REGION Network 256
   RUNG wire#powerrail
      Contact( "EMS".Carrier[41].SDC_OUT.Faults.MotionOnFault )
      Coil( "Carrier_41_Motion_On_Fault" )
   END_RUNG
   // the same network as SCL:
   "Carrier_41_Motion_On_Fault" := "EMS".Carrier[41].SDC_OUT.Faults.MotionOnFault;
END_REGION

REGION Network 257
   RUNG wire#powerrail
      Contact( "EMS".Carrier[41].SDC_OUT.Faults.MotionOffFault )
      Coil( "Carrier_41_Motion_Off_Fault" )
   END_RUNG
   // the same network as SCL:
   "Carrier_41_Motion_Off_Fault" := "EMS".Carrier[41].SDC_OUT.Faults.MotionOffFault;
END_REGION

REGION Network 258
   RUNG wire#powerrail
      Contact( "EMS".Carrier[41].SDC_OUT.Faults.CarrierSpacingFault )
      Coil( "Carrier_41_Carrier_Spacing_Fault" )
   END_RUNG
   // the same network as SCL:
   "Carrier_41_Carrier_Spacing_Fault" := "EMS".Carrier[41].SDC_OUT.Faults.CarrierSpacingFault;
END_REGION

REGION Network 259
   RUNG wire#powerrail
      Move(in := "EMS".Carrier[42].SDC_OUT.Zone, out1 => "Carrier_42_Carrier_In_Zone")
   END_RUNG
   // the same network as SCL:
   "Carrier_42_Carrier_In_Zone" := "EMS".Carrier[42].SDC_OUT.Zone;
END_REGION

REGION Network 260
   RUNG wire#powerrail
      Move(in := "EMS".Carrier[42].SDC_OUT.CarrierNum, out1 => "Carrier_42_Carrier_Number_Echo")
   END_RUNG
   // the same network as SCL:
   "Carrier_42_Carrier_Number_Echo" := "EMS".Carrier[42].SDC_OUT.CarrierNum;
END_REGION

REGION Network 261
   RUNG wire#powerrail
      Move(in := "EMS".Carrier[42].SDC_OUT.CarrierPosition, out1 => "Carrier_42_Carrier_Position_Echo")
   END_RUNG
   // the same network as SCL:
   "Carrier_42_Carrier_Position_Echo" := "EMS".Carrier[42].SDC_OUT.CarrierPosition;
END_REGION

REGION Network 262
   RUNG wire#powerrail
      Move(in := "EMS".Carrier[42].SDC_OUT.NextCarrierNum, out1 => "Carrier_42_Next_Carrier_Number")
   END_RUNG
   // the same network as SCL:
   "Carrier_42_Next_Carrier_Number" := "EMS".Carrier[42].SDC_OUT.NextCarrierNum;
END_REGION

REGION Network 263
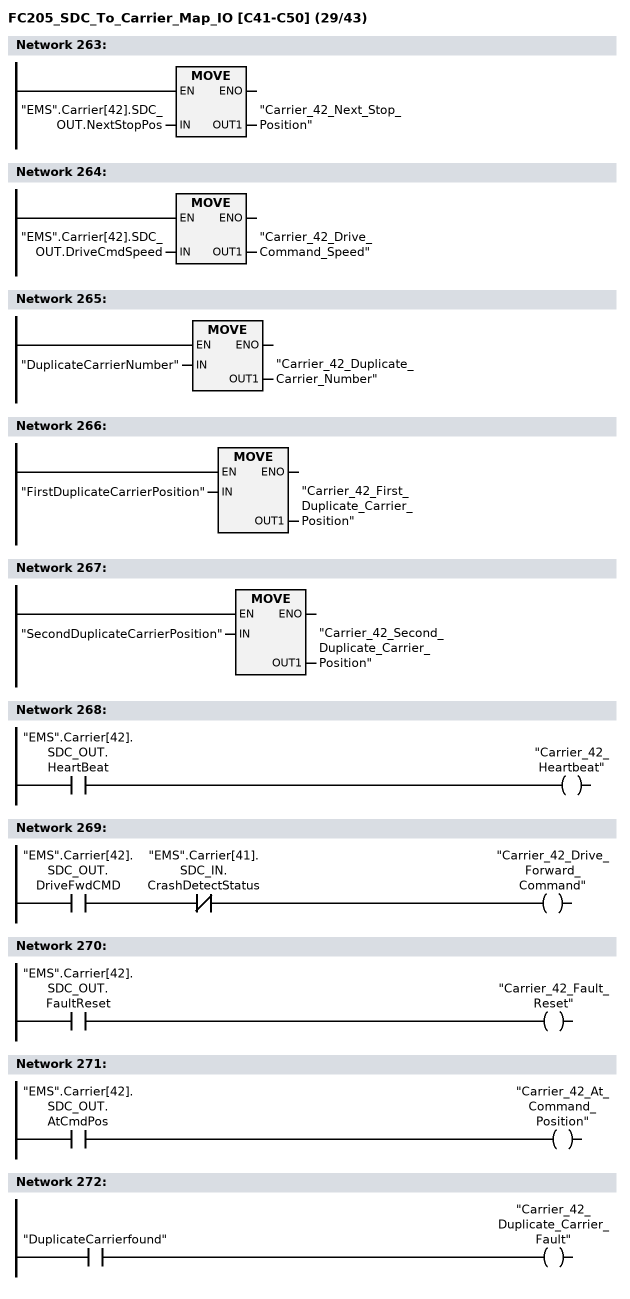
   RUNG wire#powerrail
      Move(in := "EMS".Carrier[42].SDC_OUT.NextStopPos, out1 => "Carrier_42_Next_Stop_Position")
   END_RUNG
   // the same network as SCL:
   "Carrier_42_Next_Stop_Position" := "EMS".Carrier[42].SDC_OUT.NextStopPos;
END_REGION

REGION Network 264
   RUNG wire#powerrail
      Move(in := "EMS".Carrier[42].SDC_OUT.DriveCmdSpeed, out1 => "Carrier_42_Drive_Command_Speed")
   END_RUNG
   // the same network as SCL:
   "Carrier_42_Drive_Command_Speed" := "EMS".Carrier[42].SDC_OUT.DriveCmdSpeed;
END_REGION

REGION Network 265
   RUNG wire#powerrail
      Move(in := "DuplicateCarrierNumber", out1 => "Carrier_42_Duplicate_Carrier_Number")
   END_RUNG
   // the same network as SCL:
   "Carrier_42_Duplicate_Carrier_Number" := "DuplicateCarrierNumber";
END_REGION

REGION Network 266
   RUNG wire#powerrail
      Move(in := "FirstDuplicateCarrierPosition", out1 => "Carrier_42_First_Duplicate_Carrier_Position")
   END_RUNG
   // the same network as SCL:
   "Carrier_42_First_Duplicate_Carrier_Position" := "FirstDuplicateCarrierPosition";
END_REGION

REGION Network 267
   RUNG wire#powerrail
      Move(in := "SecondDuplicateCarrierPosition", out1 => "Carrier_42_Second_Duplicate_Carrier_Position")
   END_RUNG
   // the same network as SCL:
   "Carrier_42_Second_Duplicate_Carrier_Position" := "SecondDuplicateCarrierPosition";
END_REGION

REGION Network 268
   RUNG wire#powerrail
      Contact( "EMS".Carrier[42].SDC_OUT.HeartBeat )
      Coil( "Carrier_42_Heartbeat" )
   END_RUNG
   // the same network as SCL:
   "Carrier_42_Heartbeat" := "EMS".Carrier[42].SDC_OUT.HeartBeat;
END_REGION

REGION Network 269
   RUNG wire#powerrail
      Contact( "EMS".Carrier[42].SDC_OUT.DriveFwdCMD )
      I_Contact( "EMS".Carrier[41].SDC_IN.CrashDetectStatus )
      Coil( "Carrier_42_Drive_Forward_Command" )
   END_RUNG
   // the same network as SCL:
   "Carrier_42_Drive_Forward_Command" := "EMS".Carrier[42].SDC_OUT.DriveFwdCMD AND NOT "EMS".Carrier[41].SDC_IN.CrashDetectStatus;
END_REGION

REGION Network 270
   RUNG wire#powerrail
      Contact( "EMS".Carrier[42].SDC_OUT.FaultReset )
      Coil( "Carrier_42_Fault_Reset" )
   END_RUNG
   // the same network as SCL:
   "Carrier_42_Fault_Reset" := "EMS".Carrier[42].SDC_OUT.FaultReset;
END_REGION

REGION Network 271
   RUNG wire#powerrail
      Contact( "EMS".Carrier[42].SDC_OUT.AtCmdPos )
      Coil( "Carrier_42_At_Command_Position" )
   END_RUNG
   // the same network as SCL:
   "Carrier_42_At_Command_Position" := "EMS".Carrier[42].SDC_OUT.AtCmdPos;
END_REGION

REGION Network 272
   RUNG wire#powerrail
      Contact( "DuplicateCarrierfound" )
      Coil( "Carrier_42_Duplicate_Carrier_Fault" )
   END_RUNG
   // the same network as SCL:
   "Carrier_42_Duplicate_Carrier_Fault" := "DuplicateCarrierfound";
END_REGION

REGION Network 273
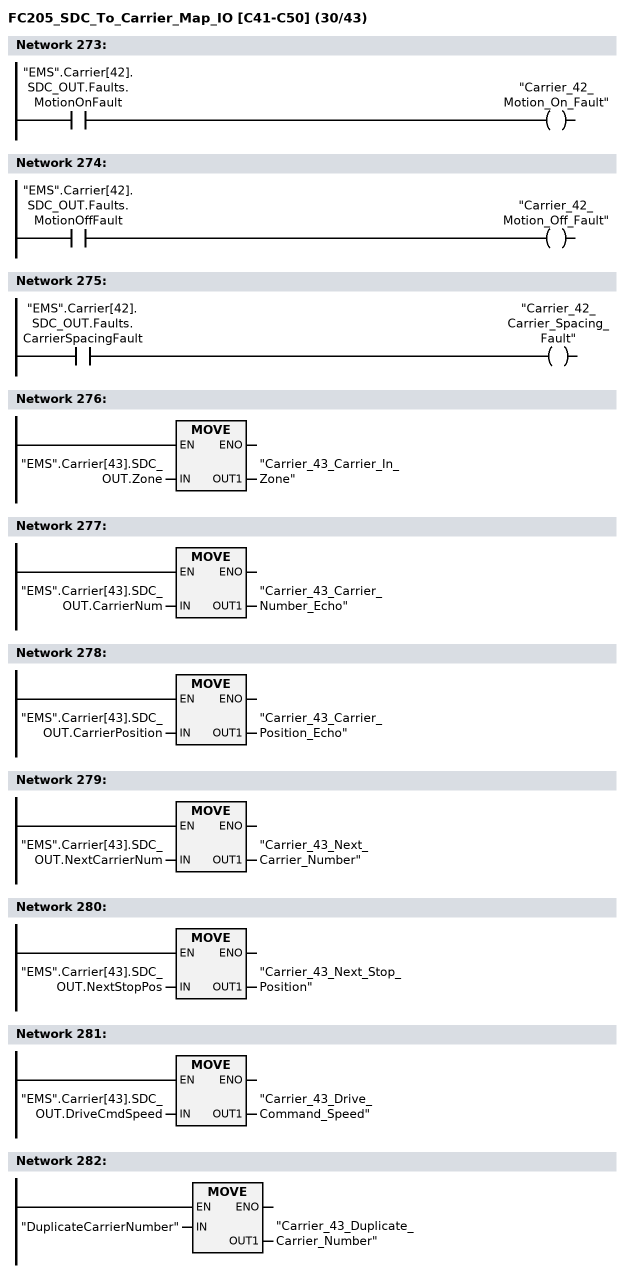
   RUNG wire#powerrail
      Contact( "EMS".Carrier[42].SDC_OUT.Faults.MotionOnFault )
      Coil( "Carrier_42_Motion_On_Fault" )
   END_RUNG
   // the same network as SCL:
   "Carrier_42_Motion_On_Fault" := "EMS".Carrier[42].SDC_OUT.Faults.MotionOnFault;
END_REGION

REGION Network 274
   RUNG wire#powerrail
      Contact( "EMS".Carrier[42].SDC_OUT.Faults.MotionOffFault )
      Coil( "Carrier_42_Motion_Off_Fault" )
   END_RUNG
   // the same network as SCL:
   "Carrier_42_Motion_Off_Fault" := "EMS".Carrier[42].SDC_OUT.Faults.MotionOffFault;
END_REGION

REGION Network 275
   RUNG wire#powerrail
      Contact( "EMS".Carrier[42].SDC_OUT.Faults.CarrierSpacingFault )
      Coil( "Carrier_42_Carrier_Spacing_Fault" )
   END_RUNG
   // the same network as SCL:
   "Carrier_42_Carrier_Spacing_Fault" := "EMS".Carrier[42].SDC_OUT.Faults.CarrierSpacingFault;
END_REGION

REGION Network 276
   RUNG wire#powerrail
      Move(in := "EMS".Carrier[43].SDC_OUT.Zone, out1 => "Carrier_43_Carrier_In_Zone")
   END_RUNG
   // the same network as SCL:
   "Carrier_43_Carrier_In_Zone" := "EMS".Carrier[43].SDC_OUT.Zone;
END_REGION

REGION Network 277
   RUNG wire#powerrail
      Move(in := "EMS".Carrier[43].SDC_OUT.CarrierNum, out1 => "Carrier_43_Carrier_Number_Echo")
   END_RUNG
   // the same network as SCL:
   "Carrier_43_Carrier_Number_Echo" := "EMS".Carrier[43].SDC_OUT.CarrierNum;
END_REGION

REGION Network 278
   RUNG wire#powerrail
      Move(in := "EMS".Carrier[43].SDC_OUT.CarrierPosition, out1 => "Carrier_43_Carrier_Position_Echo")
   END_RUNG
   // the same network as SCL:
   "Carrier_43_Carrier_Position_Echo" := "EMS".Carrier[43].SDC_OUT.CarrierPosition;
END_REGION

REGION Network 279
   RUNG wire#powerrail
      Move(in := "EMS".Carrier[43].SDC_OUT.NextCarrierNum, out1 => "Carrier_43_Next_Carrier_Number")
   END_RUNG
   // the same network as SCL:
   "Carrier_43_Next_Carrier_Number" := "EMS".Carrier[43].SDC_OUT.NextCarrierNum;
END_REGION

REGION Network 280
   RUNG wire#powerrail
      Move(in := "EMS".Carrier[43].SDC_OUT.NextStopPos, out1 => "Carrier_43_Next_Stop_Position")
   END_RUNG
   // the same network as SCL:
   "Carrier_43_Next_Stop_Position" := "EMS".Carrier[43].SDC_OUT.NextStopPos;
END_REGION

REGION Network 281
   RUNG wire#powerrail
      Move(in := "EMS".Carrier[43].SDC_OUT.DriveCmdSpeed, out1 => "Carrier_43_Drive_Command_Speed")
   END_RUNG
   // the same network as SCL:
   "Carrier_43_Drive_Command_Speed" := "EMS".Carrier[43].SDC_OUT.DriveCmdSpeed;
END_REGION

REGION Network 282
   RUNG wire#powerrail
      Move(in := "DuplicateCarrierNumber", out1 => "Carrier_43_Duplicate_Carrier_Number")
   END_RUNG
   // the same network as SCL:
   "Carrier_43_Duplicate_Carrier_Number" := "DuplicateCarrierNumber";
END_REGION

REGION Network 283
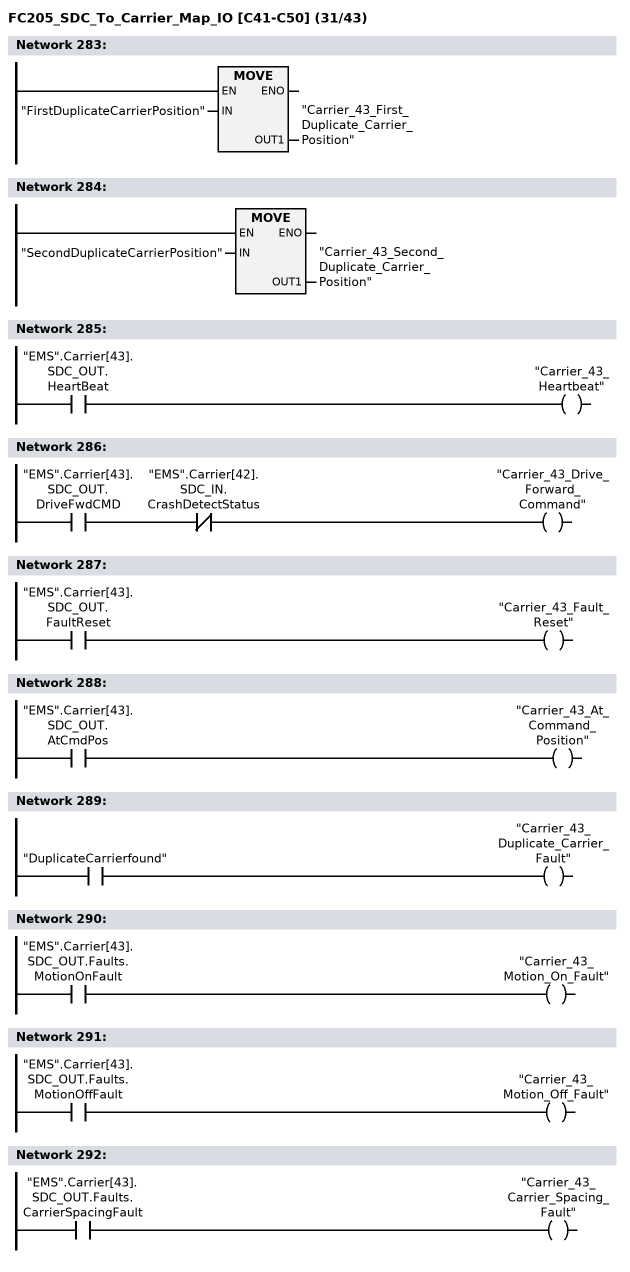
   RUNG wire#powerrail
      Move(in := "FirstDuplicateCarrierPosition", out1 => "Carrier_43_First_Duplicate_Carrier_Position")
   END_RUNG
   // the same network as SCL:
   "Carrier_43_First_Duplicate_Carrier_Position" := "FirstDuplicateCarrierPosition";
END_REGION

REGION Network 284
   RUNG wire#powerrail
      Move(in := "SecondDuplicateCarrierPosition", out1 => "Carrier_43_Second_Duplicate_Carrier_Position")
   END_RUNG
   // the same network as SCL:
   "Carrier_43_Second_Duplicate_Carrier_Position" := "SecondDuplicateCarrierPosition";
END_REGION

REGION Network 285
   RUNG wire#powerrail
      Contact( "EMS".Carrier[43].SDC_OUT.HeartBeat )
      Coil( "Carrier_43_Heartbeat" )
   END_RUNG
   // the same network as SCL:
   "Carrier_43_Heartbeat" := "EMS".Carrier[43].SDC_OUT.HeartBeat;
END_REGION

REGION Network 286
   RUNG wire#powerrail
      Contact( "EMS".Carrier[43].SDC_OUT.DriveFwdCMD )
      I_Contact( "EMS".Carrier[42].SDC_IN.CrashDetectStatus )
      Coil( "Carrier_43_Drive_Forward_Command" )
   END_RUNG
   // the same network as SCL:
   "Carrier_43_Drive_Forward_Command" := "EMS".Carrier[43].SDC_OUT.DriveFwdCMD AND NOT "EMS".Carrier[42].SDC_IN.CrashDetectStatus;
END_REGION

REGION Network 287
   RUNG wire#powerrail
      Contact( "EMS".Carrier[43].SDC_OUT.FaultReset )
      Coil( "Carrier_43_Fault_Reset" )
   END_RUNG
   // the same network as SCL:
   "Carrier_43_Fault_Reset" := "EMS".Carrier[43].SDC_OUT.FaultReset;
END_REGION

REGION Network 288
   RUNG wire#powerrail
      Contact( "EMS".Carrier[43].SDC_OUT.AtCmdPos )
      Coil( "Carrier_43_At_Command_Position" )
   END_RUNG
   // the same network as SCL:
   "Carrier_43_At_Command_Position" := "EMS".Carrier[43].SDC_OUT.AtCmdPos;
END_REGION

REGION Network 289
   RUNG wire#powerrail
      Contact( "DuplicateCarrierfound" )
      Coil( "Carrier_43_Duplicate_Carrier_Fault" )
   END_RUNG
   // the same network as SCL:
   "Carrier_43_Duplicate_Carrier_Fault" := "DuplicateCarrierfound";
END_REGION

REGION Network 290
   RUNG wire#powerrail
      Contact( "EMS".Carrier[43].SDC_OUT.Faults.MotionOnFault )
      Coil( "Carrier_43_Motion_On_Fault" )
   END_RUNG
   // the same network as SCL:
   "Carrier_43_Motion_On_Fault" := "EMS".Carrier[43].SDC_OUT.Faults.MotionOnFault;
END_REGION

REGION Network 291
   RUNG wire#powerrail
      Contact( "EMS".Carrier[43].SDC_OUT.Faults.MotionOffFault )
      Coil( "Carrier_43_Motion_Off_Fault" )
   END_RUNG
   // the same network as SCL:
   "Carrier_43_Motion_Off_Fault" := "EMS".Carrier[43].SDC_OUT.Faults.MotionOffFault;
END_REGION

REGION Network 292
   RUNG wire#powerrail
      Contact( "EMS".Carrier[43].SDC_OUT.Faults.CarrierSpacingFault )
      Coil( "Carrier_43_Carrier_Spacing_Fault" )
   END_RUNG
   // the same network as SCL:
   "Carrier_43_Carrier_Spacing_Fault" := "EMS".Carrier[43].SDC_OUT.Faults.CarrierSpacingFault;
END_REGION

REGION Network 293
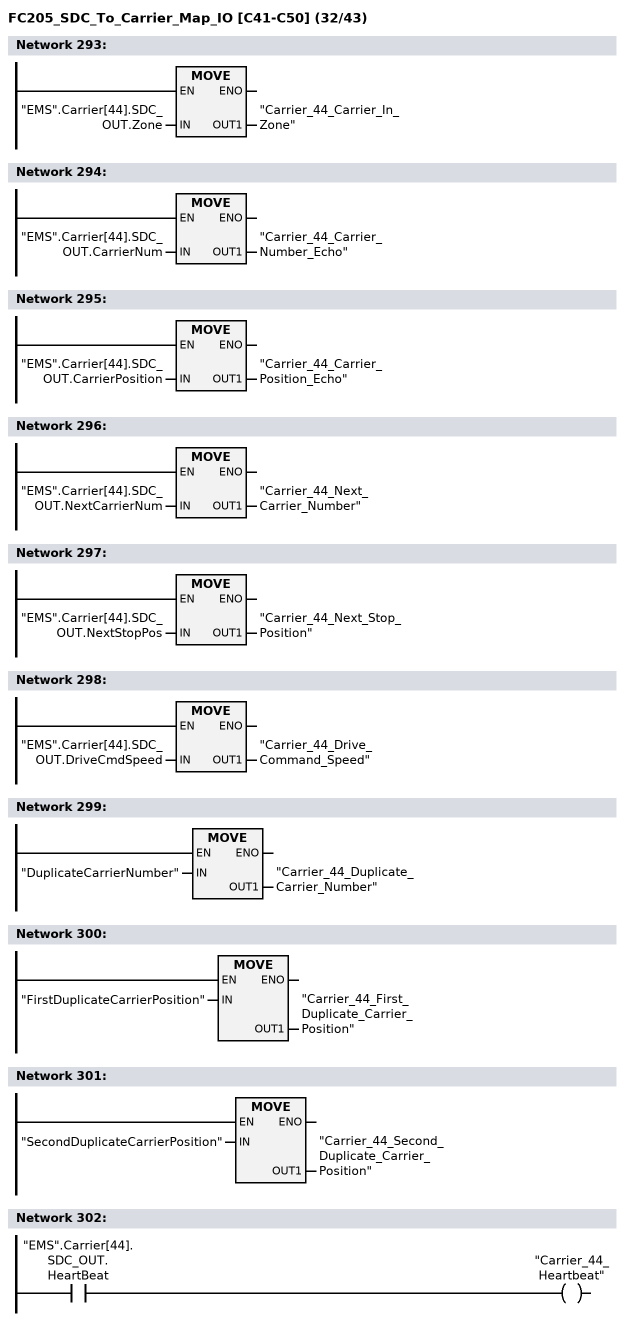
   RUNG wire#powerrail
      Move(in := "EMS".Carrier[44].SDC_OUT.Zone, out1 => "Carrier_44_Carrier_In_Zone")
   END_RUNG
   // the same network as SCL:
   "Carrier_44_Carrier_In_Zone" := "EMS".Carrier[44].SDC_OUT.Zone;
END_REGION

REGION Network 294
   RUNG wire#powerrail
      Move(in := "EMS".Carrier[44].SDC_OUT.CarrierNum, out1 => "Carrier_44_Carrier_Number_Echo")
   END_RUNG
   // the same network as SCL:
   "Carrier_44_Carrier_Number_Echo" := "EMS".Carrier[44].SDC_OUT.CarrierNum;
END_REGION

REGION Network 295
   RUNG wire#powerrail
      Move(in := "EMS".Carrier[44].SDC_OUT.CarrierPosition, out1 => "Carrier_44_Carrier_Position_Echo")
   END_RUNG
   // the same network as SCL:
   "Carrier_44_Carrier_Position_Echo" := "EMS".Carrier[44].SDC_OUT.CarrierPosition;
END_REGION

REGION Network 296
   RUNG wire#powerrail
      Move(in := "EMS".Carrier[44].SDC_OUT.NextCarrierNum, out1 => "Carrier_44_Next_Carrier_Number")
   END_RUNG
   // the same network as SCL:
   "Carrier_44_Next_Carrier_Number" := "EMS".Carrier[44].SDC_OUT.NextCarrierNum;
END_REGION

REGION Network 297
   RUNG wire#powerrail
      Move(in := "EMS".Carrier[44].SDC_OUT.NextStopPos, out1 => "Carrier_44_Next_Stop_Position")
   END_RUNG
   // the same network as SCL:
   "Carrier_44_Next_Stop_Position" := "EMS".Carrier[44].SDC_OUT.NextStopPos;
END_REGION

REGION Network 298
   RUNG wire#powerrail
      Move(in := "EMS".Carrier[44].SDC_OUT.DriveCmdSpeed, out1 => "Carrier_44_Drive_Command_Speed")
   END_RUNG
   // the same network as SCL:
   "Carrier_44_Drive_Command_Speed" := "EMS".Carrier[44].SDC_OUT.DriveCmdSpeed;
END_REGION

REGION Network 299
   RUNG wire#powerrail
      Move(in := "DuplicateCarrierNumber", out1 => "Carrier_44_Duplicate_Carrier_Number")
   END_RUNG
   // the same network as SCL:
   "Carrier_44_Duplicate_Carrier_Number" := "DuplicateCarrierNumber";
END_REGION

REGION Network 300
   RUNG wire#powerrail
      Move(in := "FirstDuplicateCarrierPosition", out1 => "Carrier_44_First_Duplicate_Carrier_Position")
   END_RUNG
   // the same network as SCL:
   "Carrier_44_First_Duplicate_Carrier_Position" := "FirstDuplicateCarrierPosition";
END_REGION

REGION Network 301
   RUNG wire#powerrail
      Move(in := "SecondDuplicateCarrierPosition", out1 => "Carrier_44_Second_Duplicate_Carrier_Position")
   END_RUNG
   // the same network as SCL:
   "Carrier_44_Second_Duplicate_Carrier_Position" := "SecondDuplicateCarrierPosition";
END_REGION

REGION Network 302
   RUNG wire#powerrail
      Contact( "EMS".Carrier[44].SDC_OUT.HeartBeat )
      Coil( "Carrier_44_Heartbeat" )
   END_RUNG
   // the same network as SCL:
   "Carrier_44_Heartbeat" := "EMS".Carrier[44].SDC_OUT.HeartBeat;
END_REGION

REGION Network 303
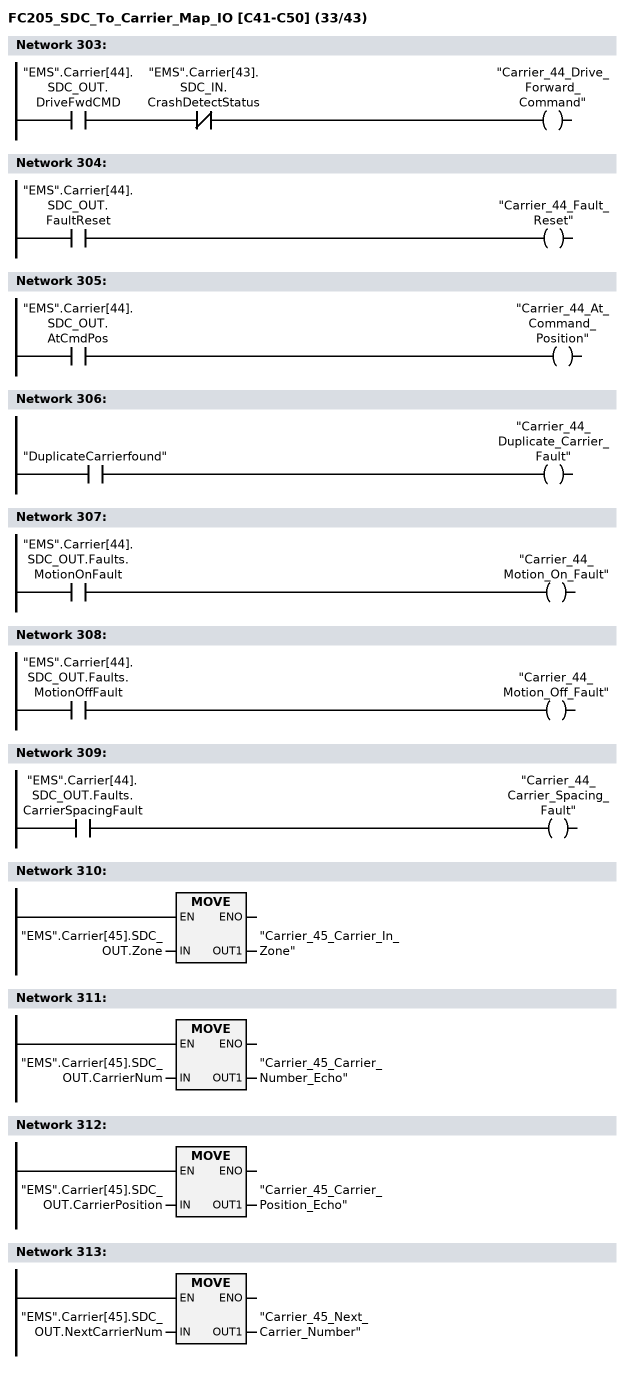
   RUNG wire#powerrail
      Contact( "EMS".Carrier[44].SDC_OUT.DriveFwdCMD )
      I_Contact( "EMS".Carrier[43].SDC_IN.CrashDetectStatus )
      Coil( "Carrier_44_Drive_Forward_Command" )
   END_RUNG
   // the same network as SCL:
   "Carrier_44_Drive_Forward_Command" := "EMS".Carrier[44].SDC_OUT.DriveFwdCMD AND NOT "EMS".Carrier[43].SDC_IN.CrashDetectStatus;
END_REGION

REGION Network 304
   RUNG wire#powerrail
      Contact( "EMS".Carrier[44].SDC_OUT.FaultReset )
      Coil( "Carrier_44_Fault_Reset" )
   END_RUNG
   // the same network as SCL:
   "Carrier_44_Fault_Reset" := "EMS".Carrier[44].SDC_OUT.FaultReset;
END_REGION

REGION Network 305
   RUNG wire#powerrail
      Contact( "EMS".Carrier[44].SDC_OUT.AtCmdPos )
      Coil( "Carrier_44_At_Command_Position" )
   END_RUNG
   // the same network as SCL:
   "Carrier_44_At_Command_Position" := "EMS".Carrier[44].SDC_OUT.AtCmdPos;
END_REGION

REGION Network 306
   RUNG wire#powerrail
      Contact( "DuplicateCarrierfound" )
      Coil( "Carrier_44_Duplicate_Carrier_Fault" )
   END_RUNG
   // the same network as SCL:
   "Carrier_44_Duplicate_Carrier_Fault" := "DuplicateCarrierfound";
END_REGION

REGION Network 307
   RUNG wire#powerrail
      Contact( "EMS".Carrier[44].SDC_OUT.Faults.MotionOnFault )
      Coil( "Carrier_44_Motion_On_Fault" )
   END_RUNG
   // the same network as SCL:
   "Carrier_44_Motion_On_Fault" := "EMS".Carrier[44].SDC_OUT.Faults.MotionOnFault;
END_REGION

REGION Network 308
   RUNG wire#powerrail
      Contact( "EMS".Carrier[44].SDC_OUT.Faults.MotionOffFault )
      Coil( "Carrier_44_Motion_Off_Fault" )
   END_RUNG
   // the same network as SCL:
   "Carrier_44_Motion_Off_Fault" := "EMS".Carrier[44].SDC_OUT.Faults.MotionOffFault;
END_REGION

REGION Network 309
   RUNG wire#powerrail
      Contact( "EMS".Carrier[44].SDC_OUT.Faults.CarrierSpacingFault )
      Coil( "Carrier_44_Carrier_Spacing_Fault" )
   END_RUNG
   // the same network as SCL:
   "Carrier_44_Carrier_Spacing_Fault" := "EMS".Carrier[44].SDC_OUT.Faults.CarrierSpacingFault;
END_REGION

REGION Network 310
   RUNG wire#powerrail
      Move(in := "EMS".Carrier[45].SDC_OUT.Zone, out1 => "Carrier_45_Carrier_In_Zone")
   END_RUNG
   // the same network as SCL:
   "Carrier_45_Carrier_In_Zone" := "EMS".Carrier[45].SDC_OUT.Zone;
END_REGION

REGION Network 311
   RUNG wire#powerrail
      Move(in := "EMS".Carrier[45].SDC_OUT.CarrierNum, out1 => "Carrier_45_Carrier_Number_Echo")
   END_RUNG
   // the same network as SCL:
   "Carrier_45_Carrier_Number_Echo" := "EMS".Carrier[45].SDC_OUT.CarrierNum;
END_REGION

REGION Network 312
   RUNG wire#powerrail
      Move(in := "EMS".Carrier[45].SDC_OUT.CarrierPosition, out1 => "Carrier_45_Carrier_Position_Echo")
   END_RUNG
   // the same network as SCL:
   "Carrier_45_Carrier_Position_Echo" := "EMS".Carrier[45].SDC_OUT.CarrierPosition;
END_REGION

REGION Network 313
   RUNG wire#powerrail
      Move(in := "EMS".Carrier[45].SDC_OUT.NextCarrierNum, out1 => "Carrier_45_Next_Carrier_Number")
   END_RUNG
   // the same network as SCL:
   "Carrier_45_Next_Carrier_Number" := "EMS".Carrier[45].SDC_OUT.NextCarrierNum;
END_REGION

REGION Network 314
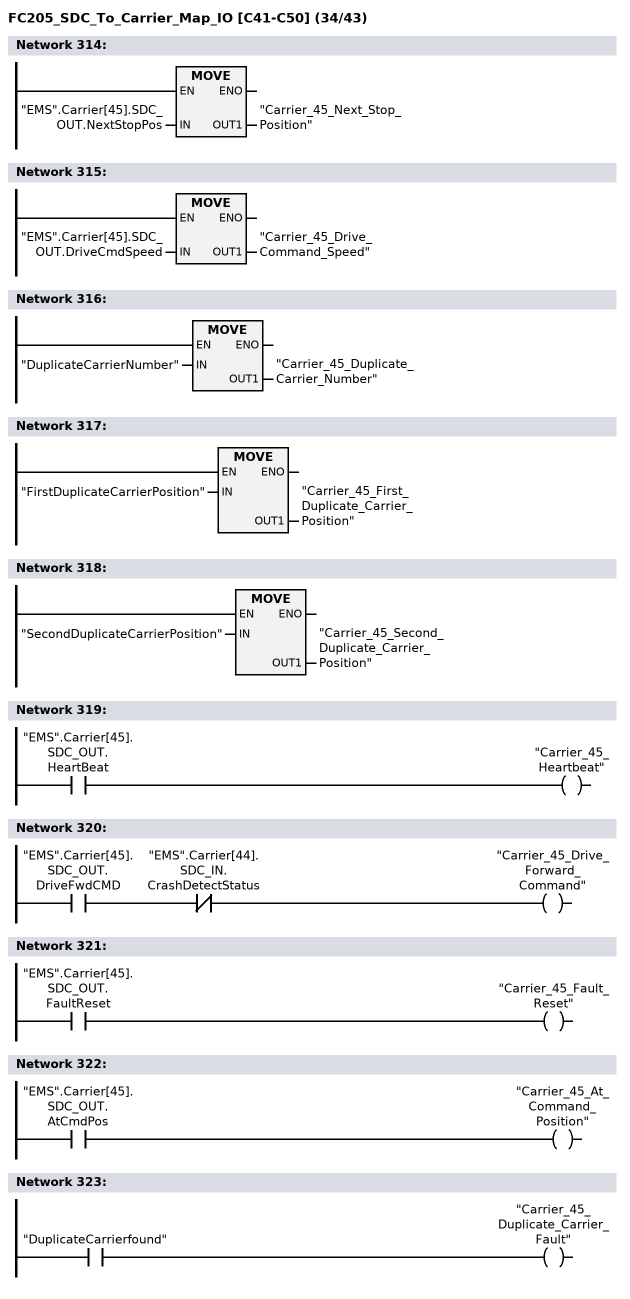
   RUNG wire#powerrail
      Move(in := "EMS".Carrier[45].SDC_OUT.NextStopPos, out1 => "Carrier_45_Next_Stop_Position")
   END_RUNG
   // the same network as SCL:
   "Carrier_45_Next_Stop_Position" := "EMS".Carrier[45].SDC_OUT.NextStopPos;
END_REGION

REGION Network 315
   RUNG wire#powerrail
      Move(in := "EMS".Carrier[45].SDC_OUT.DriveCmdSpeed, out1 => "Carrier_45_Drive_Command_Speed")
   END_RUNG
   // the same network as SCL:
   "Carrier_45_Drive_Command_Speed" := "EMS".Carrier[45].SDC_OUT.DriveCmdSpeed;
END_REGION

REGION Network 316
   RUNG wire#powerrail
      Move(in := "DuplicateCarrierNumber", out1 => "Carrier_45_Duplicate_Carrier_Number")
   END_RUNG
   // the same network as SCL:
   "Carrier_45_Duplicate_Carrier_Number" := "DuplicateCarrierNumber";
END_REGION

REGION Network 317
   RUNG wire#powerrail
      Move(in := "FirstDuplicateCarrierPosition", out1 => "Carrier_45_First_Duplicate_Carrier_Position")
   END_RUNG
   // the same network as SCL:
   "Carrier_45_First_Duplicate_Carrier_Position" := "FirstDuplicateCarrierPosition";
END_REGION

REGION Network 318
   RUNG wire#powerrail
      Move(in := "SecondDuplicateCarrierPosition", out1 => "Carrier_45_Second_Duplicate_Carrier_Position")
   END_RUNG
   // the same network as SCL:
   "Carrier_45_Second_Duplicate_Carrier_Position" := "SecondDuplicateCarrierPosition";
END_REGION

REGION Network 319
   RUNG wire#powerrail
      Contact( "EMS".Carrier[45].SDC_OUT.HeartBeat )
      Coil( "Carrier_45_Heartbeat" )
   END_RUNG
   // the same network as SCL:
   "Carrier_45_Heartbeat" := "EMS".Carrier[45].SDC_OUT.HeartBeat;
END_REGION

REGION Network 320
   RUNG wire#powerrail
      Contact( "EMS".Carrier[45].SDC_OUT.DriveFwdCMD )
      I_Contact( "EMS".Carrier[44].SDC_IN.CrashDetectStatus )
      Coil( "Carrier_45_Drive_Forward_Command" )
   END_RUNG
   // the same network as SCL:
   "Carrier_45_Drive_Forward_Command" := "EMS".Carrier[45].SDC_OUT.DriveFwdCMD AND NOT "EMS".Carrier[44].SDC_IN.CrashDetectStatus;
END_REGION

REGION Network 321
   RUNG wire#powerrail
      Contact( "EMS".Carrier[45].SDC_OUT.FaultReset )
      Coil( "Carrier_45_Fault_Reset" )
   END_RUNG
   // the same network as SCL:
   "Carrier_45_Fault_Reset" := "EMS".Carrier[45].SDC_OUT.FaultReset;
END_REGION

REGION Network 322
   RUNG wire#powerrail
      Contact( "EMS".Carrier[45].SDC_OUT.AtCmdPos )
      Coil( "Carrier_45_At_Command_Position" )
   END_RUNG
   // the same network as SCL:
   "Carrier_45_At_Command_Position" := "EMS".Carrier[45].SDC_OUT.AtCmdPos;
END_REGION

REGION Network 323
   RUNG wire#powerrail
      Contact( "DuplicateCarrierfound" )
      Coil( "Carrier_45_Duplicate_Carrier_Fault" )
   END_RUNG
   // the same network as SCL:
   "Carrier_45_Duplicate_Carrier_Fault" := "DuplicateCarrierfound";
END_REGION

REGION Network 324
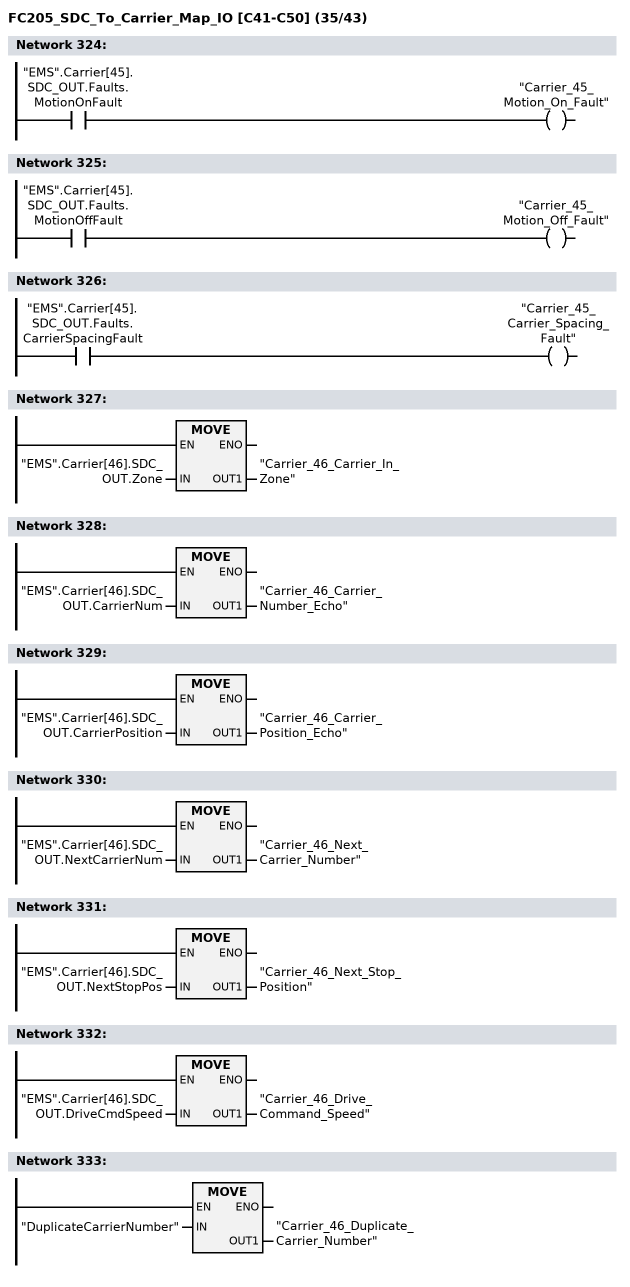
   RUNG wire#powerrail
      Contact( "EMS".Carrier[45].SDC_OUT.Faults.MotionOnFault )
      Coil( "Carrier_45_Motion_On_Fault" )
   END_RUNG
   // the same network as SCL:
   "Carrier_45_Motion_On_Fault" := "EMS".Carrier[45].SDC_OUT.Faults.MotionOnFault;
END_REGION

REGION Network 325
   RUNG wire#powerrail
      Contact( "EMS".Carrier[45].SDC_OUT.Faults.MotionOffFault )
      Coil( "Carrier_45_Motion_Off_Fault" )
   END_RUNG
   // the same network as SCL:
   "Carrier_45_Motion_Off_Fault" := "EMS".Carrier[45].SDC_OUT.Faults.MotionOffFault;
END_REGION

REGION Network 326
   RUNG wire#powerrail
      Contact( "EMS".Carrier[45].SDC_OUT.Faults.CarrierSpacingFault )
      Coil( "Carrier_45_Carrier_Spacing_Fault" )
   END_RUNG
   // the same network as SCL:
   "Carrier_45_Carrier_Spacing_Fault" := "EMS".Carrier[45].SDC_OUT.Faults.CarrierSpacingFault;
END_REGION

REGION Network 327
   RUNG wire#powerrail
      Move(in := "EMS".Carrier[46].SDC_OUT.Zone, out1 => "Carrier_46_Carrier_In_Zone")
   END_RUNG
   // the same network as SCL:
   "Carrier_46_Carrier_In_Zone" := "EMS".Carrier[46].SDC_OUT.Zone;
END_REGION

REGION Network 328
   RUNG wire#powerrail
      Move(in := "EMS".Carrier[46].SDC_OUT.CarrierNum, out1 => "Carrier_46_Carrier_Number_Echo")
   END_RUNG
   // the same network as SCL:
   "Carrier_46_Carrier_Number_Echo" := "EMS".Carrier[46].SDC_OUT.CarrierNum;
END_REGION

REGION Network 329
   RUNG wire#powerrail
      Move(in := "EMS".Carrier[46].SDC_OUT.CarrierPosition, out1 => "Carrier_46_Carrier_Position_Echo")
   END_RUNG
   // the same network as SCL:
   "Carrier_46_Carrier_Position_Echo" := "EMS".Carrier[46].SDC_OUT.CarrierPosition;
END_REGION

REGION Network 330
   RUNG wire#powerrail
      Move(in := "EMS".Carrier[46].SDC_OUT.NextCarrierNum, out1 => "Carrier_46_Next_Carrier_Number")
   END_RUNG
   // the same network as SCL:
   "Carrier_46_Next_Carrier_Number" := "EMS".Carrier[46].SDC_OUT.NextCarrierNum;
END_REGION

REGION Network 331
   RUNG wire#powerrail
      Move(in := "EMS".Carrier[46].SDC_OUT.NextStopPos, out1 => "Carrier_46_Next_Stop_Position")
   END_RUNG
   // the same network as SCL:
   "Carrier_46_Next_Stop_Position" := "EMS".Carrier[46].SDC_OUT.NextStopPos;
END_REGION

REGION Network 332
   RUNG wire#powerrail
      Move(in := "EMS".Carrier[46].SDC_OUT.DriveCmdSpeed, out1 => "Carrier_46_Drive_Command_Speed")
   END_RUNG
   // the same network as SCL:
   "Carrier_46_Drive_Command_Speed" := "EMS".Carrier[46].SDC_OUT.DriveCmdSpeed;
END_REGION

REGION Network 333
   RUNG wire#powerrail
      Move(in := "DuplicateCarrierNumber", out1 => "Carrier_46_Duplicate_Carrier_Number")
   END_RUNG
   // the same network as SCL:
   "Carrier_46_Duplicate_Carrier_Number" := "DuplicateCarrierNumber";
END_REGION

REGION Network 334
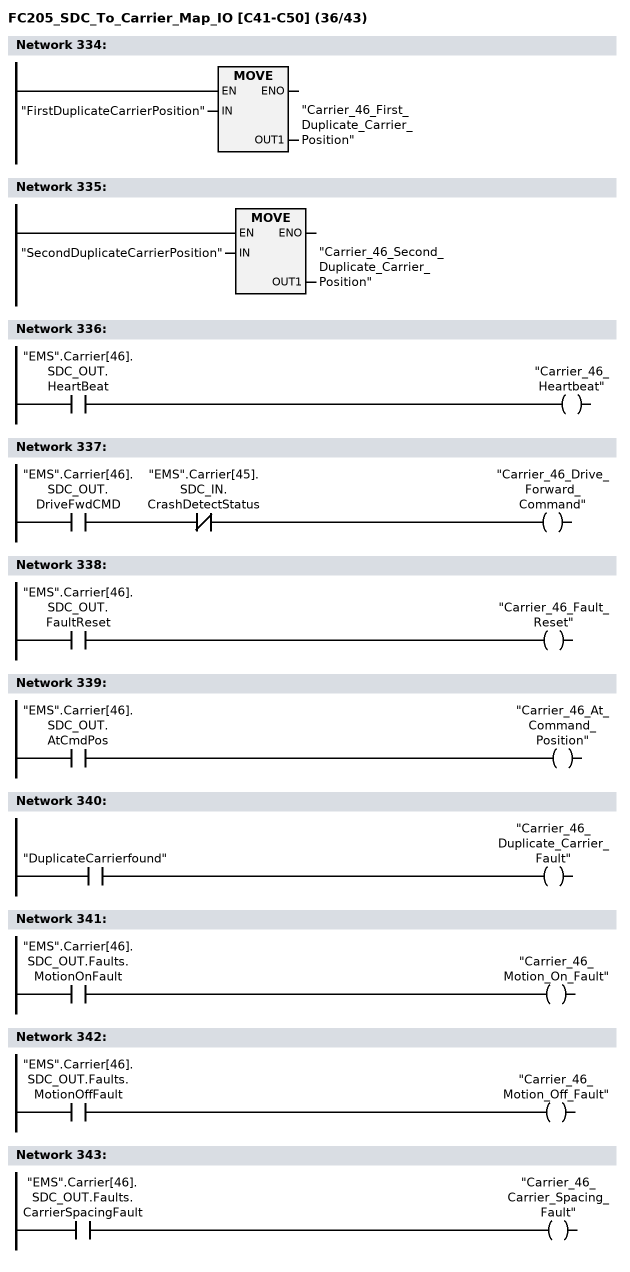
   RUNG wire#powerrail
      Move(in := "FirstDuplicateCarrierPosition", out1 => "Carrier_46_First_Duplicate_Carrier_Position")
   END_RUNG
   // the same network as SCL:
   "Carrier_46_First_Duplicate_Carrier_Position" := "FirstDuplicateCarrierPosition";
END_REGION

REGION Network 335
   RUNG wire#powerrail
      Move(in := "SecondDuplicateCarrierPosition", out1 => "Carrier_46_Second_Duplicate_Carrier_Position")
   END_RUNG
   // the same network as SCL:
   "Carrier_46_Second_Duplicate_Carrier_Position" := "SecondDuplicateCarrierPosition";
END_REGION

REGION Network 336
   RUNG wire#powerrail
      Contact( "EMS".Carrier[46].SDC_OUT.HeartBeat )
      Coil( "Carrier_46_Heartbeat" )
   END_RUNG
   // the same network as SCL:
   "Carrier_46_Heartbeat" := "EMS".Carrier[46].SDC_OUT.HeartBeat;
END_REGION

REGION Network 337
   RUNG wire#powerrail
      Contact( "EMS".Carrier[46].SDC_OUT.DriveFwdCMD )
      I_Contact( "EMS".Carrier[45].SDC_IN.CrashDetectStatus )
      Coil( "Carrier_46_Drive_Forward_Command" )
   END_RUNG
   // the same network as SCL:
   "Carrier_46_Drive_Forward_Command" := "EMS".Carrier[46].SDC_OUT.DriveFwdCMD AND NOT "EMS".Carrier[45].SDC_IN.CrashDetectStatus;
END_REGION

REGION Network 338
   RUNG wire#powerrail
      Contact( "EMS".Carrier[46].SDC_OUT.FaultReset )
      Coil( "Carrier_46_Fault_Reset" )
   END_RUNG
   // the same network as SCL:
   "Carrier_46_Fault_Reset" := "EMS".Carrier[46].SDC_OUT.FaultReset;
END_REGION

REGION Network 339
   RUNG wire#powerrail
      Contact( "EMS".Carrier[46].SDC_OUT.AtCmdPos )
      Coil( "Carrier_46_At_Command_Position" )
   END_RUNG
   // the same network as SCL:
   "Carrier_46_At_Command_Position" := "EMS".Carrier[46].SDC_OUT.AtCmdPos;
END_REGION

REGION Network 340
   RUNG wire#powerrail
      Contact( "DuplicateCarrierfound" )
      Coil( "Carrier_46_Duplicate_Carrier_Fault" )
   END_RUNG
   // the same network as SCL:
   "Carrier_46_Duplicate_Carrier_Fault" := "DuplicateCarrierfound";
END_REGION

REGION Network 341
   RUNG wire#powerrail
      Contact( "EMS".Carrier[46].SDC_OUT.Faults.MotionOnFault )
      Coil( "Carrier_46_Motion_On_Fault" )
   END_RUNG
   // the same network as SCL:
   "Carrier_46_Motion_On_Fault" := "EMS".Carrier[46].SDC_OUT.Faults.MotionOnFault;
END_REGION

REGION Network 342
   RUNG wire#powerrail
      Contact( "EMS".Carrier[46].SDC_OUT.Faults.MotionOffFault )
      Coil( "Carrier_46_Motion_Off_Fault" )
   END_RUNG
   // the same network as SCL:
   "Carrier_46_Motion_Off_Fault" := "EMS".Carrier[46].SDC_OUT.Faults.MotionOffFault;
END_REGION
